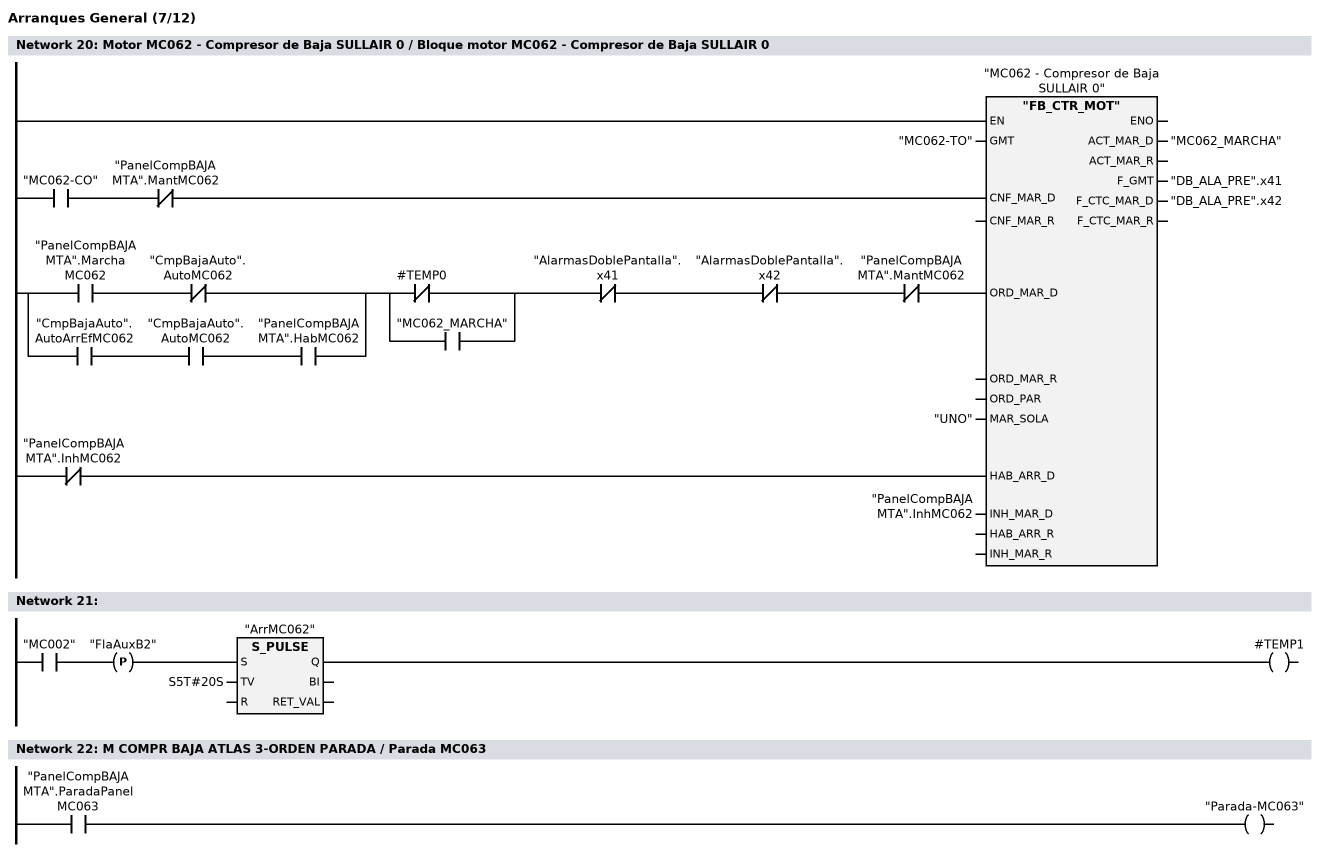
   RUNG wire#powerrail
      "MC062 - Compresor de Baja SULLAIR 0"(CNF_MAR_D := wire#w1, ORD_MAR_D := wire#w4, HAB_ARR_D := wire#w5, GMT := "MC062-TO", CNF_MAR_R :=, ORD_MAR_R :=, ORD_PAR :=, MAR_SOLA := "UNO", INH_MAR_D := "PanelCompBAJA MTA".InhMC062, HAB_ARR_R :=, INH_MAR_R :=, ACT_MAR_D => "MC062_MARCHA", ACT_MAR_R =>, F_GMT => "DB_ALA_PRE".x41, F_CTC_MAR_D => "DB_ALA_PRE".x42, F_CTC_MAR_R =>)
   END_RUNG
   RUNG wire#powerrail
      Contact( "MC062-CO" )
      I_Contact( "PanelCompBAJA MTA".MantMC062 )
   END_RUNG wire#w1
   RUNG wire#powerrail
      Contact( "PanelCompBAJA MTA".MarchaMC062 )
      I_Contact( "CmpBajaAuto".AutoMC062 )
      wire#w2
      I_Contact( #TEMP0 )
      wire#w3
      I_Contact( "AlarmasDoblePantalla".x41 )
      I_Contact( "AlarmasDoblePantalla".x42 )
      I_Contact( "PanelCompBAJA MTA".MantMC062 )
   END_RUNG wire#w4
   RUNG wire#powerrail
      Contact( "CmpBajaAuto".AutoArrEfMC062 )
      Contact( "CmpBajaAuto".AutoMC062 )
      Contact( "PanelCompBAJA MTA".HabMC062 )
   END_RUNG wire#w2
   RUNG wire#w2
      Contact( "MC062_MARCHA" )
   END_RUNG wire#w3
   RUNG wire#powerrail
      I_Contact( "PanelCompBAJA MTA".InhMC062 )
   END_RUNG wire#w5
   // the same network as SCL:
   "MC062 - Compresor de Baja SULLAIR 0"(GMT := "MC062-TO",   // "FB_CTR_MOT"
                           CNF_MAR_D := "MC062-CO" AND NOT "PanelCompBAJA MTA".MantMC062,
                           ORD_MAR_D := (("PanelCompBAJA MTA".MarchaMC062 AND NOT "CmpBajaAuto".AutoMC062) OR ("CmpBajaAuto".AutoArrEfMC062 AND "CmpBajaAuto".AutoMC062 AND "PanelCompBAJA MTA".HabMC062)) AND (NOT #TEMP0 OR "MC062_MARCHA") AND NOT "AlarmasDoblePantalla".x41 AND NOT "AlarmasDoblePantalla".x42 AND NOT "PanelCompBAJA MTA".MantMC062,
                           MAR_SOLA := "UNO",
                           HAB_ARR_D := NOT "PanelCompBAJA MTA".InhMC062,
                           INH_MAR_D := "PanelCompBAJA MTA".InhMC062,
                           ACT_MAR_D => "MC062_MARCHA",
                           F_GMT => "DB_ALA_PRE".x41,
                           F_CTC_MAR_D => "DB_ALA_PRE".x42);
END_REGION

REGION Network 21
   RUNG wire#powerrail
      Contact( "MC002" )
      P_Trig( "FlaAuxB2" )
      S_PULSE(T_NO := "ArrMC062", TV := S5T#20S, R :=, BI =>, RET_VAL =>)
      Coil( #TEMP1 )
   END_RUNG
   // the same network as SCL:
   #_w1 := "MC002" AND NOT "FlaAuxB2";   // rising edge
   "FlaAuxB2" := "MC002";
   #_s5time1 := S_PULSE(T_NO := "ArrMC062", S := #_w1, TV := S5T#20S, Q => #_w2);
   #TEMP1 := #_w2;
END_REGION

REGION Network 22: M COMPR BAJA ATLAS 3-ORDEN PARADA / Parada MC063
   RUNG wire#powerrail
      Contact( "PanelCompBAJA MTA".ParadaPanelMC063 )
      Coil( "Parada-MC063" )
   END_RUNG
   // the same network as SCL:
   "Parada-MC063" := "PanelCompBAJA MTA".ParadaPanelMC063;
END_REGION

REGION Network 23: Motor MC063 - Compresor de Baja ATLAS 3 / Bloque motor MC063 - Compresor de Baja ATLAS 3
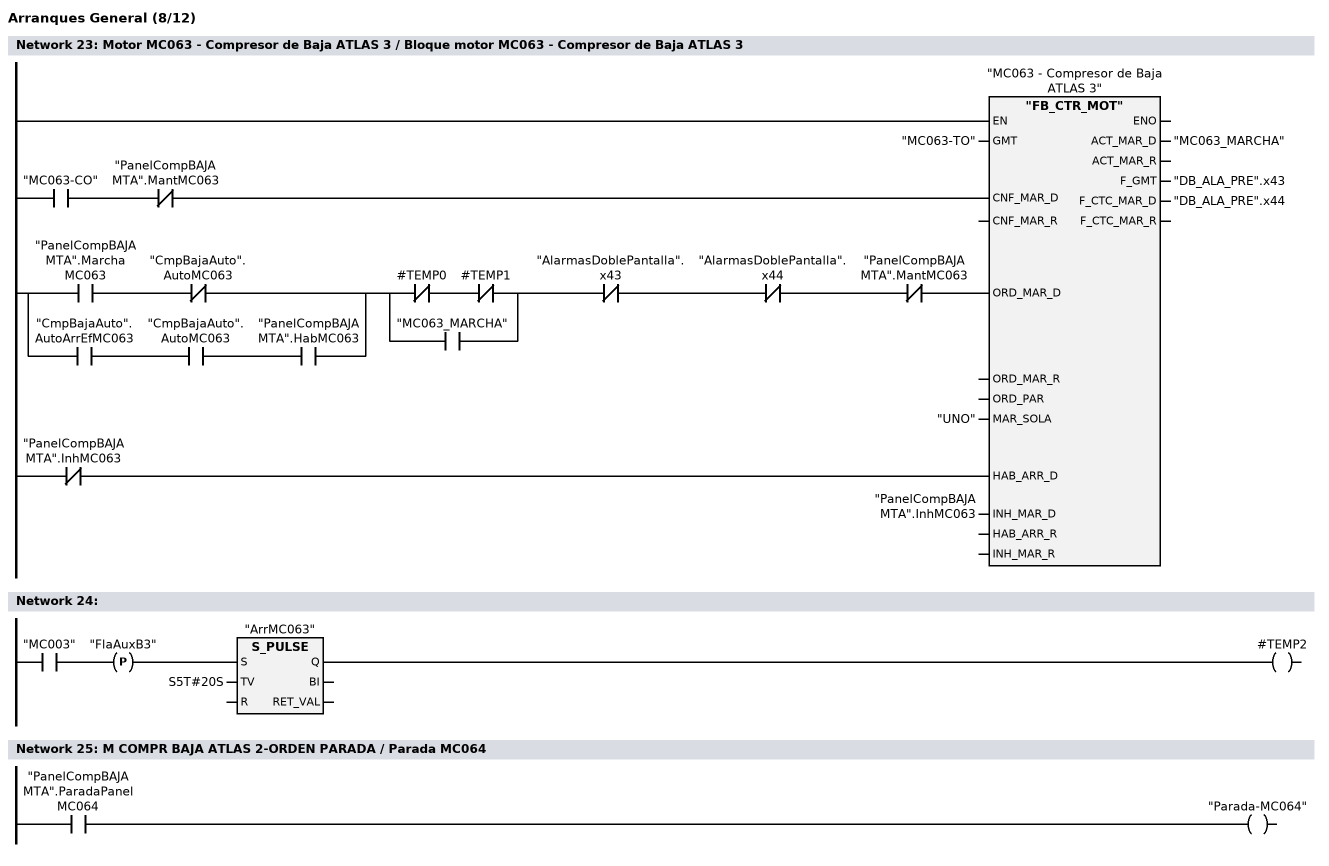
   RUNG wire#powerrail
      "MC063 - Compresor de Baja ATLAS 3"(GMT := "MC063-TO", CNF_MAR_R :=, ORD_MAR_R :=, ORD_PAR :=, MAR_SOLA := "UNO", INH_MAR_D := "PanelCompBAJA MTA".InhMC063, HAB_ARR_R :=, INH_MAR_R :=, ACT_MAR_D => "MC063_MARCHA", ACT_MAR_R =>, F_GMT => "DB_ALA_PRE".x43, F_CTC_MAR_D => "DB_ALA_PRE".x44, F_CTC_MAR_R =>, CNF_MAR_D := wire#w1, ORD_MAR_D := wire#w4, HAB_ARR_D := wire#w5)
   END_RUNG
   RUNG wire#powerrail
      Contact( "MC063-CO" )
      I_Contact( "PanelCompBAJA MTA".MantMC063 )
   END_RUNG wire#w1
   RUNG wire#powerrail
      Contact( "PanelCompBAJA MTA".MarchaMC063 )
      I_Contact( "CmpBajaAuto".AutoMC063 )
      wire#w2
      I_Contact( #TEMP0 )
      I_Contact( #TEMP1 )
      wire#w3
      I_Contact( "AlarmasDoblePantalla".x43 )
      I_Contact( "AlarmasDoblePantalla".x44 )
      I_Contact( "PanelCompBAJA MTA".MantMC063 )
   END_RUNG wire#w4
   RUNG wire#powerrail
      Contact( "CmpBajaAuto".AutoArrEfMC063 )
      Contact( "CmpBajaAuto".AutoMC063 )
      Contact( "PanelCompBAJA MTA".HabMC063 )
   END_RUNG wire#w2
   RUNG wire#w2
      Contact( "MC063_MARCHA" )
   END_RUNG wire#w3
   RUNG wire#powerrail
      I_Contact( "PanelCompBAJA MTA".InhMC063 )
   END_RUNG wire#w5
   // the same network as SCL:
   "MC063 - Compresor de Baja ATLAS 3"(GMT := "MC063-TO",   // "FB_CTR_MOT"
                           CNF_MAR_D := "MC063-CO" AND NOT "PanelCompBAJA MTA".MantMC063,
                           ORD_MAR_D := (("PanelCompBAJA MTA".MarchaMC063 AND NOT "CmpBajaAuto".AutoMC063) OR ("CmpBajaAuto".AutoArrEfMC063 AND "CmpBajaAuto".AutoMC063 AND "PanelCompBAJA MTA".HabMC063)) AND ((NOT #TEMP0 AND NOT #TEMP1) OR "MC063_MARCHA") AND NOT "AlarmasDoblePantalla".x43 AND NOT "AlarmasDoblePantalla".x44 AND NOT "PanelCompBAJA MTA".MantMC063,
                           MAR_SOLA := "UNO",
                           HAB_ARR_D := NOT "PanelCompBAJA MTA".InhMC063,
                           INH_MAR_D := "PanelCompBAJA MTA".InhMC063,
                           ACT_MAR_D => "MC063_MARCHA",
                           F_GMT => "DB_ALA_PRE".x43,
                           F_CTC_MAR_D => "DB_ALA_PRE".x44);
END_REGION

REGION Network 24
   RUNG wire#powerrail
      Contact( "MC003" )
      P_Trig( "FlaAuxB3" )
      S_PULSE(T_NO := "ArrMC063", TV := S5T#20S, R :=, BI =>, RET_VAL =>)
      Coil( #TEMP2 )
   END_RUNG
   // the same network as SCL:
   #_w1 := "MC003" AND NOT "FlaAuxB3";   // rising edge
   "FlaAuxB3" := "MC003";
   #_s5time1 := S_PULSE(T_NO := "ArrMC063", S := #_w1, TV := S5T#20S, Q => #_w2);
   #TEMP2 := #_w2;
END_REGION

REGION Network 25: M COMPR BAJA ATLAS 2-ORDEN PARADA / Parada MC064
   RUNG wire#powerrail
      Contact( "PanelCompBAJA MTA".ParadaPanelMC064 )
      Coil( "Parada-MC064" )
   END_RUNG
   // the same network as SCL:
   "Parada-MC064" := "PanelCompBAJA MTA".ParadaPanelMC064;
END_REGION

REGION Network 26: Motor MC064 - Compresor de Baja ATLAS 2 / Bloque motor MC064 - Compresor de Baja ATLAS 2
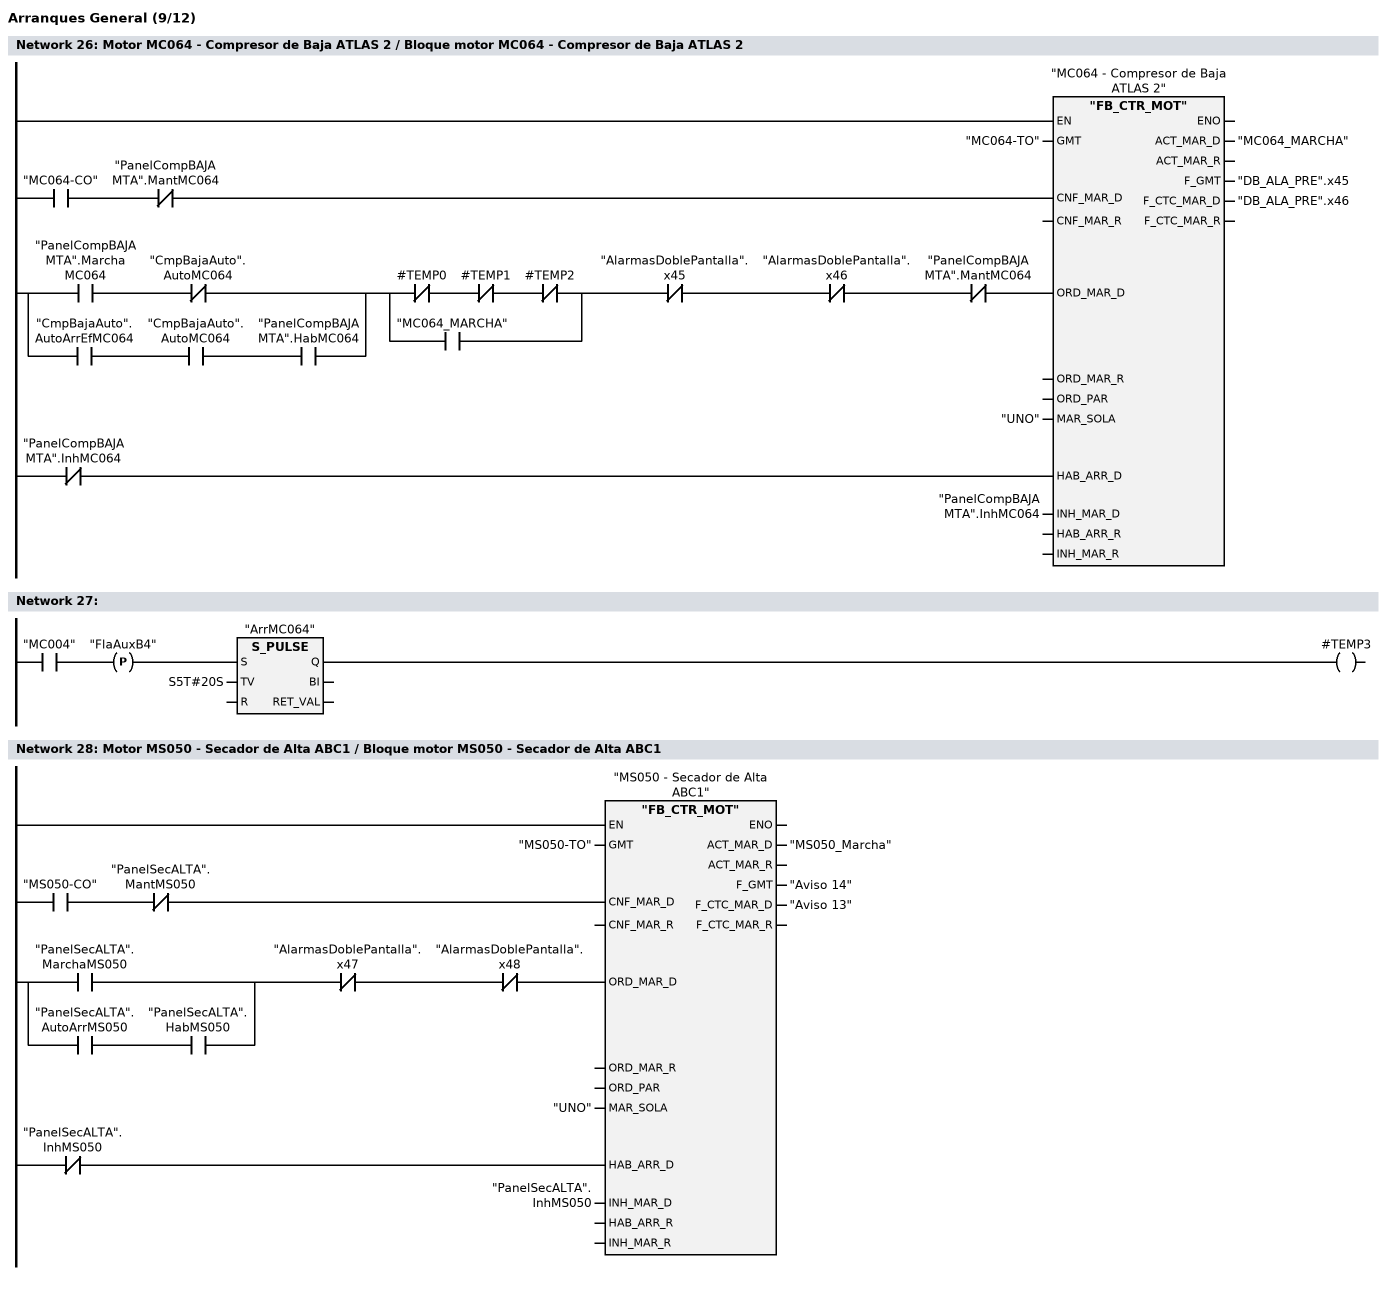
   RUNG wire#powerrail
      "MC064 - Compresor de Baja ATLAS 2"(CNF_MAR_D := wire#w1, ORD_MAR_D := wire#w4, HAB_ARR_D := wire#w5, GMT := "MC064-TO", CNF_MAR_R :=, ORD_MAR_R :=, ORD_PAR :=, MAR_SOLA := "UNO", INH_MAR_D := "PanelCompBAJA MTA".InhMC064, HAB_ARR_R :=, INH_MAR_R :=, ACT_MAR_D => "MC064_MARCHA", ACT_MAR_R =>, F_GMT => "DB_ALA_PRE".x45, F_CTC_MAR_D => "DB_ALA_PRE".x46, F_CTC_MAR_R =>)
   END_RUNG
   RUNG wire#powerrail
      Contact( "MC064-CO" )
      I_Contact( "PanelCompBAJA MTA".MantMC064 )
   END_RUNG wire#w1
   RUNG wire#powerrail
      Contact( "PanelCompBAJA MTA".MarchaMC064 )
      I_Contact( "CmpBajaAuto".AutoMC064 )
      wire#w2
      I_Contact( #TEMP0 )
      I_Contact( #TEMP1 )
      I_Contact( #TEMP2 )
      wire#w3
      I_Contact( "AlarmasDoblePantalla".x45 )
      I_Contact( "AlarmasDoblePantalla".x46 )
      I_Contact( "PanelCompBAJA MTA".MantMC064 )
   END_RUNG wire#w4
   RUNG wire#powerrail
      Contact( "CmpBajaAuto".AutoArrEfMC064 )
      Contact( "CmpBajaAuto".AutoMC064 )
      Contact( "PanelCompBAJA MTA".HabMC064 )
   END_RUNG wire#w2
   RUNG wire#w2
      Contact( "MC064_MARCHA" )
   END_RUNG wire#w3
   RUNG wire#powerrail
      I_Contact( "PanelCompBAJA MTA".InhMC064 )
   END_RUNG wire#w5
   // the same network as SCL:
   "MC064 - Compresor de Baja ATLAS 2"(GMT := "MC064-TO",   // "FB_CTR_MOT"
                           CNF_MAR_D := "MC064-CO" AND NOT "PanelCompBAJA MTA".MantMC064,
                           ORD_MAR_D := (("PanelCompBAJA MTA".MarchaMC064 AND NOT "CmpBajaAuto".AutoMC064) OR ("CmpBajaAuto".AutoArrEfMC064 AND "CmpBajaAuto".AutoMC064 AND "PanelCompBAJA MTA".HabMC064)) AND ((NOT #TEMP0 AND NOT #TEMP1 AND NOT #TEMP2) OR "MC064_MARCHA") AND NOT "AlarmasDoblePantalla".x45 AND NOT "AlarmasDoblePantalla".x46 AND NOT "PanelCompBAJA MTA".MantMC064,
                           MAR_SOLA := "UNO",
                           HAB_ARR_D := NOT "PanelCompBAJA MTA".InhMC064,
                           INH_MAR_D := "PanelCompBAJA MTA".InhMC064,
                           ACT_MAR_D => "MC064_MARCHA",
                           F_GMT => "DB_ALA_PRE".x45,
                           F_CTC_MAR_D => "DB_ALA_PRE".x46);
END_REGION

REGION Network 27
   RUNG wire#powerrail
      Contact( "MC004" )
      P_Trig( "FlaAuxB4" )
      S_PULSE(T_NO := "ArrMC064", TV := S5T#20S, R :=, BI =>, RET_VAL =>)
      Coil( #TEMP3 )
   END_RUNG
   // the same network as SCL:
   #_w1 := "MC004" AND NOT "FlaAuxB4";   // rising edge
   "FlaAuxB4" := "MC004";
   #_s5time1 := S_PULSE(T_NO := "ArrMC064", S := #_w1, TV := S5T#20S, Q => #_w2);
   #TEMP3 := #_w2;
END_REGION

REGION Network 28: Motor MS050 - Secador de Alta ABC1 / Bloque motor MS050 - Secador de Alta ABC1
   RUNG wire#powerrail
      "MS050 - Secador de Alta  ABC1"(CNF_MAR_D := wire#w1, ORD_MAR_D := wire#w3, HAB_ARR_D := wire#w4, GMT := "MS050-TO", CNF_MAR_R :=, ORD_MAR_R :=, ORD_PAR :=, MAR_SOLA := "UNO", INH_MAR_D := "PanelSecALTA".InhMS050, HAB_ARR_R :=, INH_MAR_R :=, ACT_MAR_D => "MS050_Marcha", ACT_MAR_R =>, F_GMT => "Aviso 14", F_CTC_MAR_D => "Aviso 13", F_CTC_MAR_R =>)
   END_RUNG
   RUNG wire#powerrail
      Contact( "MS050-CO" )
      I_Contact( "PanelSecALTA".MantMS050 )
   END_RUNG wire#w1
   RUNG wire#powerrail
      Contact( "PanelSecALTA".MarchaMS050 )
      wire#w2
      I_Contact( "AlarmasDoblePantalla".x47 )
      I_Contact( "AlarmasDoblePantalla".x48 )
   END_RUNG wire#w3
   RUNG wire#powerrail
      Contact( "PanelSecALTA".AutoArrMS050 )
      Contact( "PanelSecALTA".HabMS050 )
   END_RUNG wire#w2
   RUNG wire#powerrail
      I_Contact( "PanelSecALTA".InhMS050 )
   END_RUNG wire#w4
   // the same network as SCL:
   "MS050 - Secador de Alta  ABC1"(GMT := "MS050-TO",   // "FB_CTR_MOT"
                           CNF_MAR_D := "MS050-CO" AND NOT "PanelSecALTA".MantMS050,
                           ORD_MAR_D := ("PanelSecALTA".MarchaMS050 OR ("PanelSecALTA".AutoArrMS050 AND "PanelSecALTA".HabMS050)) AND NOT "AlarmasDoblePantalla".x47 AND NOT "AlarmasDoblePantalla".x48,
                           MAR_SOLA := "UNO",
                           HAB_ARR_D := NOT "PanelSecALTA".InhMS050,
                           INH_MAR_D := "PanelSecALTA".InhMS050,
                           ACT_MAR_D => "MS050_Marcha",
                           F_GMT => "Aviso 14",
                           F_CTC_MAR_D => "Aviso 13");
END_REGION

REGION Network 29: Motor MS051 - Secador de Alta ABC3 / Bloque motor MS051 - Secador de Alta ABC3
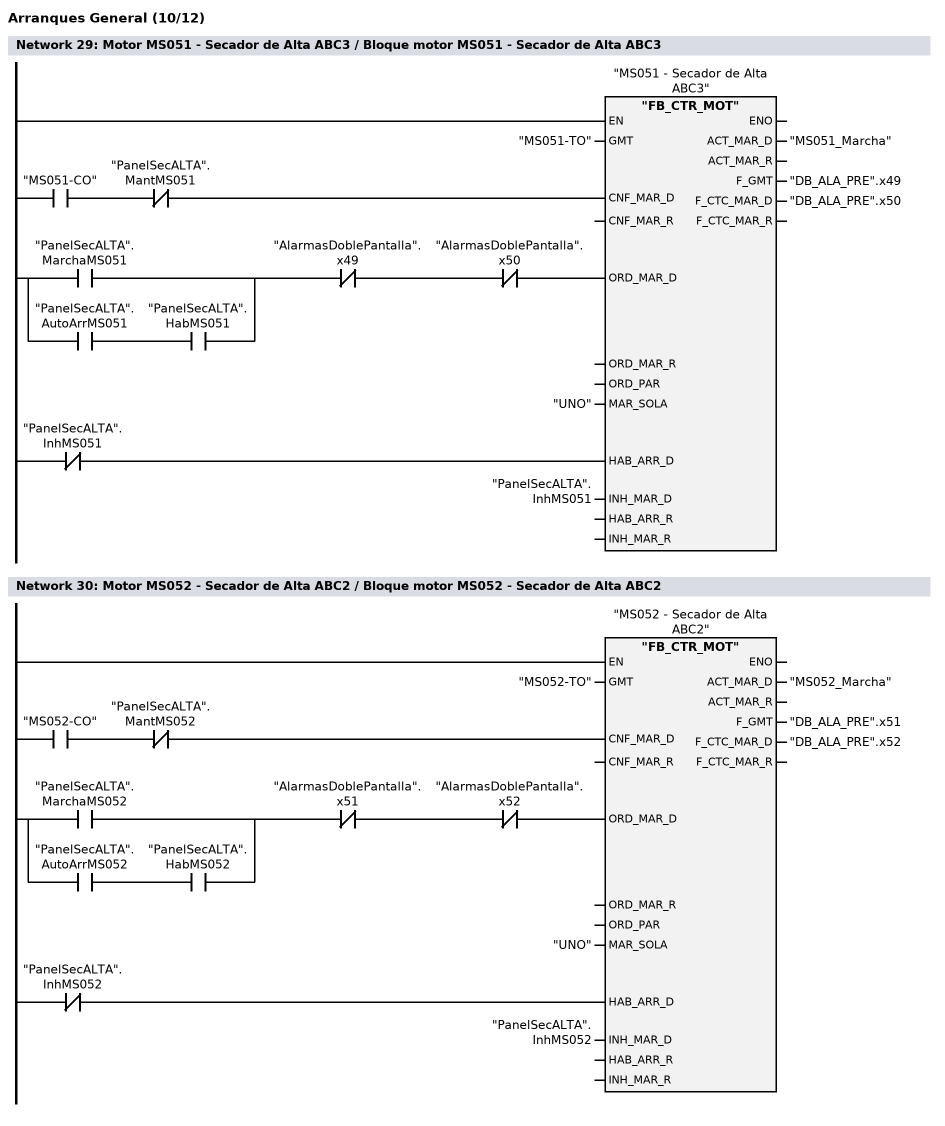
   RUNG wire#powerrail
      "MS051 - Secador de Alta  ABC3"(CNF_MAR_D := wire#w1, ORD_MAR_D := wire#w3, HAB_ARR_D := wire#w4, GMT := "MS051-TO", CNF_MAR_R :=, ORD_MAR_R :=, ORD_PAR :=, MAR_SOLA := "UNO", INH_MAR_D := "PanelSecALTA".InhMS051, HAB_ARR_R :=, INH_MAR_R :=, ACT_MAR_D => "MS051_Marcha", ACT_MAR_R =>, F_GMT => "DB_ALA_PRE".x49, F_CTC_MAR_D => "DB_ALA_PRE".x50, F_CTC_MAR_R =>)
   END_RUNG
   RUNG wire#powerrail
      Contact( "MS051-CO" )
      I_Contact( "PanelSecALTA".MantMS051 )
   END_RUNG wire#w1
   RUNG wire#powerrail
      Contact( "PanelSecALTA".MarchaMS051 )
      wire#w2
      I_Contact( "AlarmasDoblePantalla".x49 )
      I_Contact( "AlarmasDoblePantalla".x50 )
   END_RUNG wire#w3
   RUNG wire#powerrail
      Contact( "PanelSecALTA".AutoArrMS051 )
      Contact( "PanelSecALTA".HabMS051 )
   END_RUNG wire#w2
   RUNG wire#powerrail
      I_Contact( "PanelSecALTA".InhMS051 )
   END_RUNG wire#w4
   // the same network as SCL:
   "MS051 - Secador de Alta  ABC3"(GMT := "MS051-TO",   // "FB_CTR_MOT"
                           CNF_MAR_D := "MS051-CO" AND NOT "PanelSecALTA".MantMS051,
                           ORD_MAR_D := ("PanelSecALTA".MarchaMS051 OR ("PanelSecALTA".AutoArrMS051 AND "PanelSecALTA".HabMS051)) AND NOT "AlarmasDoblePantalla".x49 AND NOT "AlarmasDoblePantalla".x50,
                           MAR_SOLA := "UNO",
                           HAB_ARR_D := NOT "PanelSecALTA".InhMS051,
                           INH_MAR_D := "PanelSecALTA".InhMS051,
                           ACT_MAR_D => "MS051_Marcha",
                           F_GMT => "DB_ALA_PRE".x49,
                           F_CTC_MAR_D => "DB_ALA_PRE".x50);
END_REGION

REGION Network 30: Motor MS052 - Secador de Alta ABC2 / Bloque motor MS052 - Secador de Alta ABC2
   RUNG wire#powerrail
      "MS052 - Secador de Alta  ABC2"(CNF_MAR_D := wire#w1, ORD_MAR_D := wire#w3, HAB_ARR_D := wire#w4, GMT := "MS052-TO", CNF_MAR_R :=, ORD_MAR_R :=, ORD_PAR :=, MAR_SOLA := "UNO", INH_MAR_D := "PanelSecALTA".InhMS052, HAB_ARR_R :=, INH_MAR_R :=, ACT_MAR_D => "MS052_Marcha", ACT_MAR_R =>, F_GMT => "DB_ALA_PRE".x51, F_CTC_MAR_D => "DB_ALA_PRE".x52, F_CTC_MAR_R =>)
   END_RUNG
   RUNG wire#powerrail
      Contact( "MS052-CO" )
      I_Contact( "PanelSecALTA".MantMS052 )
   END_RUNG wire#w1
   RUNG wire#powerrail
      Contact( "PanelSecALTA".MarchaMS052 )
      wire#w2
      I_Contact( "AlarmasDoblePantalla".x51 )
      I_Contact( "AlarmasDoblePantalla".x52 )
   END_RUNG wire#w3
   RUNG wire#powerrail
      Contact( "PanelSecALTA".AutoArrMS052 )
      Contact( "PanelSecALTA".HabMS052 )
   END_RUNG wire#w2
   RUNG wire#powerrail
      I_Contact( "PanelSecALTA".InhMS052 )
   END_RUNG wire#w4
   // the same network as SCL:
   "MS052 - Secador de Alta  ABC2"(GMT := "MS052-TO",   // "FB_CTR_MOT"
                           CNF_MAR_D := "MS052-CO" AND NOT "PanelSecALTA".MantMS052,
                           ORD_MAR_D := ("PanelSecALTA".MarchaMS052 OR ("PanelSecALTA".AutoArrMS052 AND "PanelSecALTA".HabMS052)) AND NOT "AlarmasDoblePantalla".x51 AND NOT "AlarmasDoblePantalla".x52,
                           MAR_SOLA := "UNO",
                           HAB_ARR_D := NOT "PanelSecALTA".InhMS052,
                           INH_MAR_D := "PanelSecALTA".InhMS052,
                           ACT_MAR_D => "MS052_Marcha",
                           F_GMT => "DB_ALA_PRE".x51,
                           F_CTC_MAR_D => "DB_ALA_PRE".x52);
END_REGION

REGION Network 31: Motor MS053 - Secador de Alta FARGON / Bloque motor MS053 - Secador de Alta FARGON
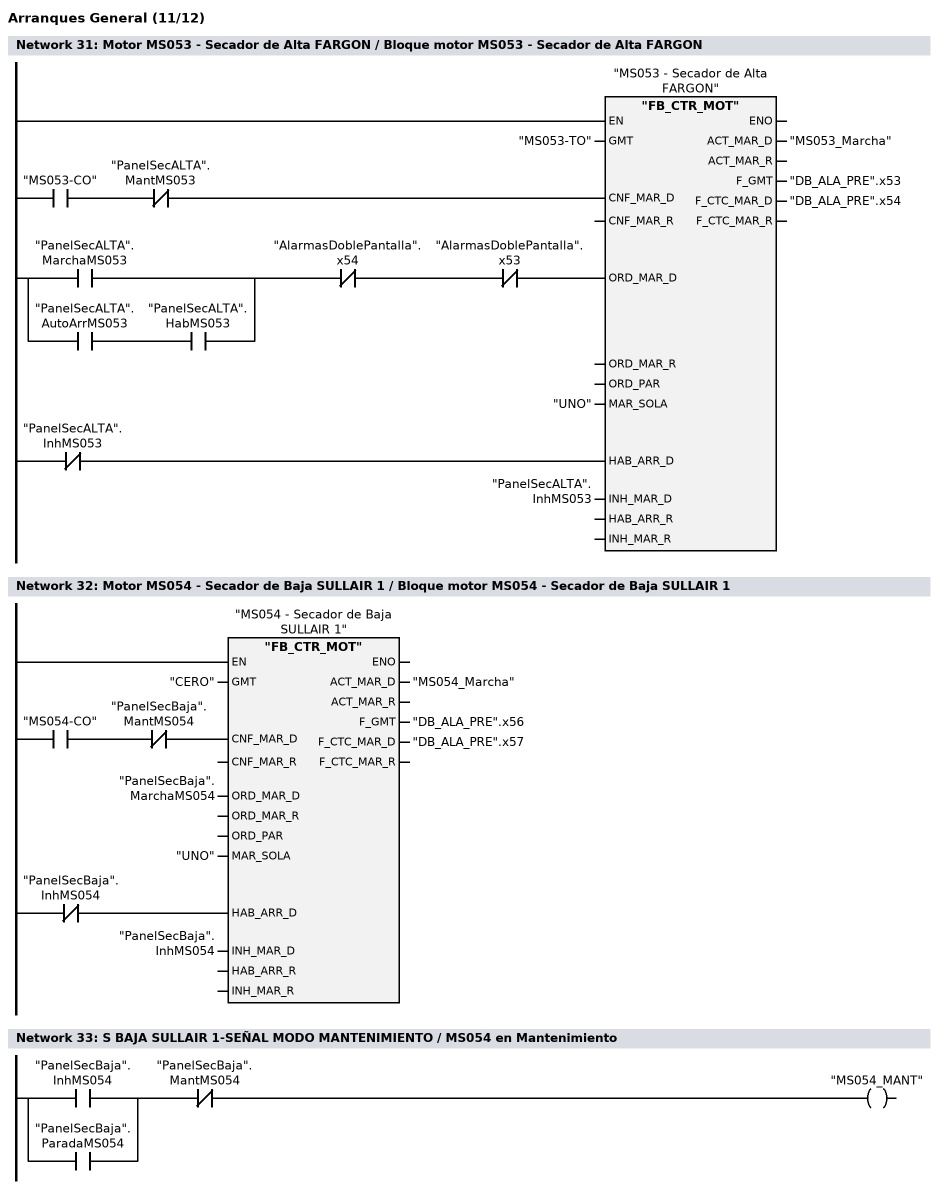
   RUNG wire#powerrail
      "MS053 - Secador de Alta  FARGON"(CNF_MAR_D := wire#w1, ORD_MAR_D := wire#w3, HAB_ARR_D := wire#w4, GMT := "MS053-TO", CNF_MAR_R :=, ORD_MAR_R :=, ORD_PAR :=, MAR_SOLA := "UNO", INH_MAR_D := "PanelSecALTA".InhMS053, HAB_ARR_R :=, INH_MAR_R :=, ACT_MAR_D => "MS053_Marcha", ACT_MAR_R =>, F_GMT => "DB_ALA_PRE".x53, F_CTC_MAR_D => "DB_ALA_PRE".x54, F_CTC_MAR_R =>)
   END_RUNG
   RUNG wire#powerrail
      Contact( "MS053-CO" )
      I_Contact( "PanelSecALTA".MantMS053 )
   END_RUNG wire#w1
   RUNG wire#powerrail
      Contact( "PanelSecALTA".MarchaMS053 )
      wire#w2
      I_Contact( "AlarmasDoblePantalla".x54 )
      I_Contact( "AlarmasDoblePantalla".x53 )
   END_RUNG wire#w3
   RUNG wire#powerrail
      Contact( "PanelSecALTA".AutoArrMS053 )
      Contact( "PanelSecALTA".HabMS053 )
   END_RUNG wire#w2
   RUNG wire#powerrail
      I_Contact( "PanelSecALTA".InhMS053 )
   END_RUNG wire#w4
   // the same network as SCL:
   "MS053 - Secador de Alta  FARGON"(GMT := "MS053-TO",   // "FB_CTR_MOT"
                           CNF_MAR_D := "MS053-CO" AND NOT "PanelSecALTA".MantMS053,
                           ORD_MAR_D := ("PanelSecALTA".MarchaMS053 OR ("PanelSecALTA".AutoArrMS053 AND "PanelSecALTA".HabMS053)) AND NOT "AlarmasDoblePantalla".x54 AND NOT "AlarmasDoblePantalla".x53,
                           MAR_SOLA := "UNO",
                           HAB_ARR_D := NOT "PanelSecALTA".InhMS053,
                           INH_MAR_D := "PanelSecALTA".InhMS053,
                           ACT_MAR_D => "MS053_Marcha",
                           F_GMT => "DB_ALA_PRE".x53,
                           F_CTC_MAR_D => "DB_ALA_PRE".x54);
END_REGION

REGION Network 32: Motor MS054 - Secador de Baja SULLAIR 1 / Bloque motor MS054 - Secador de Baja SULLAIR 1
   RUNG wire#powerrail
      "MS054 - Secador de Baja SULLAIR 1"(GMT := "CERO", CNF_MAR_R :=, ORD_MAR_D := "PanelSecBaja".MarchaMS054, ORD_MAR_R :=, ORD_PAR :=, MAR_SOLA := "UNO", INH_MAR_D := "PanelSecBaja".InhMS054, HAB_ARR_R :=, INH_MAR_R :=, ACT_MAR_D => "MS054_Marcha", ACT_MAR_R =>, F_GMT => "DB_ALA_PRE".x56, F_CTC_MAR_D => "DB_ALA_PRE".x57, F_CTC_MAR_R =>, CNF_MAR_D := wire#w1, HAB_ARR_D := wire#w2)
   END_RUNG
   RUNG wire#powerrail
      Contact( "MS054-CO" )
      I_Contact( "PanelSecBaja".MantMS054 )
   END_RUNG wire#w1
   RUNG wire#powerrail
      I_Contact( "PanelSecBaja".InhMS054 )
   END_RUNG wire#w2
   // the same network as SCL:
   "MS054 - Secador de Baja SULLAIR 1"(GMT := "CERO",   // "FB_CTR_MOT"
                           CNF_MAR_D := "MS054-CO" AND NOT "PanelSecBaja".MantMS054,
                           ORD_MAR_D := "PanelSecBaja".MarchaMS054,
                           MAR_SOLA := "UNO",
                           HAB_ARR_D := NOT "PanelSecBaja".InhMS054,
                           INH_MAR_D := "PanelSecBaja".InhMS054,
                           ACT_MAR_D => "MS054_Marcha",
                           F_GMT => "DB_ALA_PRE".x56,
                           F_CTC_MAR_D => "DB_ALA_PRE".x57);
END_REGION

REGION Network 33: S BAJA SULLAIR 1-SEÑAL MODO MANTENIMIENTO / MS054 en Mantenimiento
   RUNG wire#powerrail
      Contact( "PanelSecBaja".InhMS054 )
      wire#w1
      I_Contact( "PanelSecBaja".MantMS054 )
      Coil( "MS054_MANT" )
   END_RUNG
   RUNG wire#powerrail
      Contact( "PanelSecBaja".ParadaMS054 )
   END_RUNG wire#w1
   // the same network as SCL:
   "MS054_MANT" := ("PanelSecBaja".InhMS054 OR "PanelSecBaja".ParadaMS054) AND NOT "PanelSecBaja".MantMS054;
END_REGION

REGION Network 34: Motor MS055 / Bloque motor MS055 - Secador de Baja SULLAIR 2
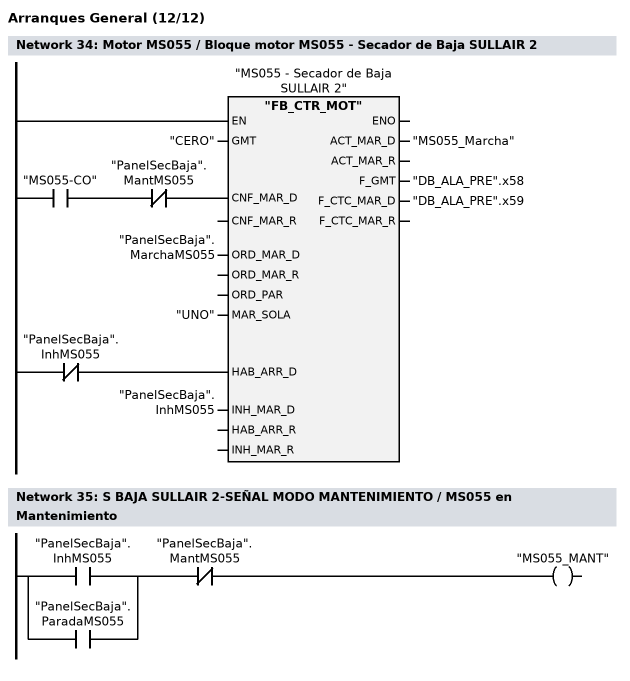
   RUNG wire#powerrail
      "MS055 - Secador de Baja SULLAIR 2"(GMT := "CERO", CNF_MAR_R :=, ORD_MAR_D := "PanelSecBaja".MarchaMS055, ORD_MAR_R :=, ORD_PAR :=, MAR_SOLA := "UNO", INH_MAR_D := "PanelSecBaja".InhMS055, HAB_ARR_R :=, INH_MAR_R :=, ACT_MAR_D => "MS055_Marcha", ACT_MAR_R =>, F_GMT => "DB_ALA_PRE".x58, F_CTC_MAR_D => "DB_ALA_PRE".x59, F_CTC_MAR_R =>, CNF_MAR_D := wire#w1, HAB_ARR_D := wire#w2)
   END_RUNG
   RUNG wire#powerrail
      Contact( "MS055-CO" )
      I_Contact( "PanelSecBaja".MantMS055 )
   END_RUNG wire#w1
   RUNG wire#powerrail
      I_Contact( "PanelSecBaja".InhMS055 )
   END_RUNG wire#w2
   // the same network as SCL:
   "MS055 - Secador de Baja SULLAIR 2"(GMT := "CERO",   // "FB_CTR_MOT"
                           CNF_MAR_D := "MS055-CO" AND NOT "PanelSecBaja".MantMS055,
                           ORD_MAR_D := "PanelSecBaja".MarchaMS055,
                           MAR_SOLA := "UNO",
                           HAB_ARR_D := NOT "PanelSecBaja".InhMS055,
                           INH_MAR_D := "PanelSecBaja".InhMS055,
                           ACT_MAR_D => "MS055_Marcha",
                           F_GMT => "DB_ALA_PRE".x58,
                           F_CTC_MAR_D => "DB_ALA_PRE".x59);
END_REGION

REGION Network 35: S BAJA SULLAIR 2-SEÑAL MODO MANTENIMIENTO / MS055 en Mantenimiento
   RUNG wire#powerrail
      Contact( "PanelSecBaja".InhMS055 )
      wire#w1
      I_Contact( "PanelSecBaja".MantMS055 )
      Coil( "MS055_MANT" )
   END_RUNG
   RUNG wire#powerrail
      Contact( "PanelSecBaja".ParadaMS055 )
   END_RUNG wire#w1
   // the same network as SCL:
   "MS055_MANT" := ("PanelSecBaja".InhMS055 OR "PanelSecBaja".ParadaMS055) AND NOT "PanelSecBaja".MantMS055;
END_REGION
END_FUNCTION
